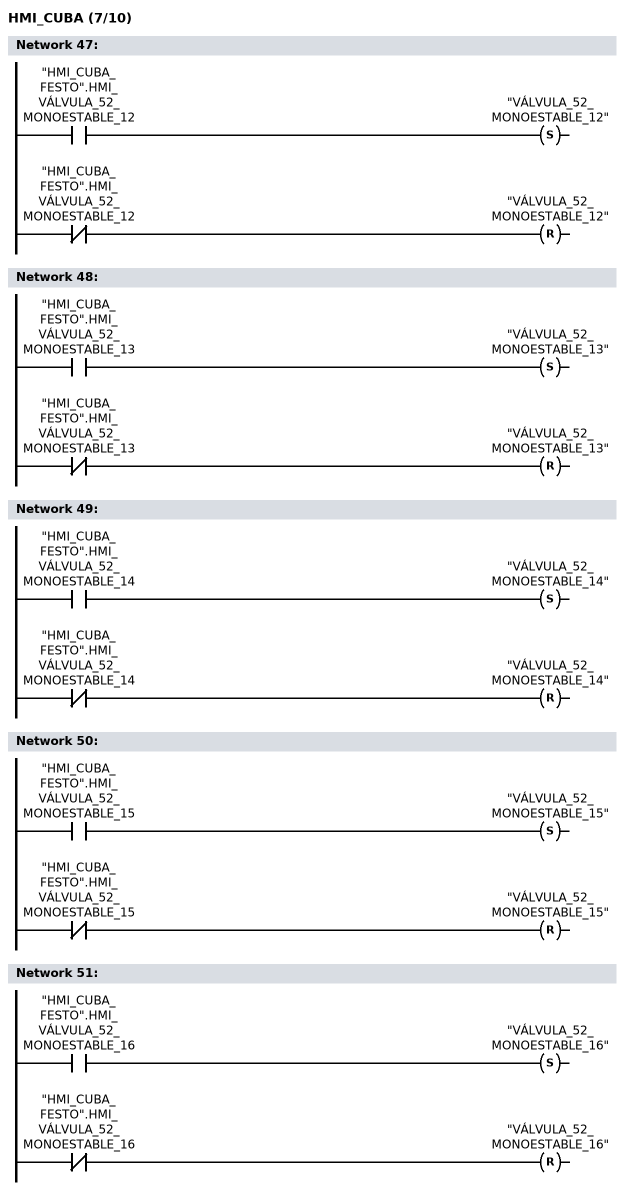
   RUNG wire#powerrail
      Contact( "HMI_CUBA_FESTO".HMI_VÁLVULA_52_MONOESTABLE_12 )
      S_Coil( "VÁLVULA_52_MONOESTABLE_12" )
   END_RUNG
   RUNG wire#powerrail
      I_Contact( "HMI_CUBA_FESTO".HMI_VÁLVULA_52_MONOESTABLE_12 )
      R_Coil( "VÁLVULA_52_MONOESTABLE_12" )
   END_RUNG
   // the same network as SCL:
   IF "HMI_CUBA_FESTO".HMI_VÁLVULA_52_MONOESTABLE_12 THEN "VÁLVULA_52_MONOESTABLE_12" := TRUE; END_IF;
   IF NOT "HMI_CUBA_FESTO".HMI_VÁLVULA_52_MONOESTABLE_12 THEN "VÁLVULA_52_MONOESTABLE_12" := FALSE; END_IF;
END_REGION

REGION Network 48
   RUNG wire#powerrail
      Contact( "HMI_CUBA_FESTO".HMI_VÁLVULA_52_MONOESTABLE_13 )
      S_Coil( "VÁLVULA_52_MONOESTABLE_13" )
   END_RUNG
   RUNG wire#powerrail
      I_Contact( "HMI_CUBA_FESTO".HMI_VÁLVULA_52_MONOESTABLE_13 )
      R_Coil( "VÁLVULA_52_MONOESTABLE_13" )
   END_RUNG
   // the same network as SCL:
   IF "HMI_CUBA_FESTO".HMI_VÁLVULA_52_MONOESTABLE_13 THEN "VÁLVULA_52_MONOESTABLE_13" := TRUE; END_IF;
   IF NOT "HMI_CUBA_FESTO".HMI_VÁLVULA_52_MONOESTABLE_13 THEN "VÁLVULA_52_MONOESTABLE_13" := FALSE; END_IF;
END_REGION

REGION Network 49
   RUNG wire#powerrail
      Contact( "HMI_CUBA_FESTO".HMI_VÁLVULA_52_MONOESTABLE_14 )
      S_Coil( "VÁLVULA_52_MONOESTABLE_14" )
   END_RUNG
   RUNG wire#powerrail
      I_Contact( "HMI_CUBA_FESTO".HMI_VÁLVULA_52_MONOESTABLE_14 )
      R_Coil( "VÁLVULA_52_MONOESTABLE_14" )
   END_RUNG
   // the same network as SCL:
   IF "HMI_CUBA_FESTO".HMI_VÁLVULA_52_MONOESTABLE_14 THEN "VÁLVULA_52_MONOESTABLE_14" := TRUE; END_IF;
   IF NOT "HMI_CUBA_FESTO".HMI_VÁLVULA_52_MONOESTABLE_14 THEN "VÁLVULA_52_MONOESTABLE_14" := FALSE; END_IF;
END_REGION

REGION Network 50
   RUNG wire#powerrail
      Contact( "HMI_CUBA_FESTO".HMI_VÁLVULA_52_MONOESTABLE_15 )
      S_Coil( "VÁLVULA_52_MONOESTABLE_15" )
   END_RUNG
   RUNG wire#powerrail
      I_Contact( "HMI_CUBA_FESTO".HMI_VÁLVULA_52_MONOESTABLE_15 )
      R_Coil( "VÁLVULA_52_MONOESTABLE_15" )
   END_RUNG
   // the same network as SCL:
   IF "HMI_CUBA_FESTO".HMI_VÁLVULA_52_MONOESTABLE_15 THEN "VÁLVULA_52_MONOESTABLE_15" := TRUE; END_IF;
   IF NOT "HMI_CUBA_FESTO".HMI_VÁLVULA_52_MONOESTABLE_15 THEN "VÁLVULA_52_MONOESTABLE_15" := FALSE; END_IF;
END_REGION

REGION Network 51
   RUNG wire#powerrail
      Contact( "HMI_CUBA_FESTO".HMI_VÁLVULA_52_MONOESTABLE_16 )
      S_Coil( "VÁLVULA_52_MONOESTABLE_16" )
   END_RUNG
   RUNG wire#powerrail
      I_Contact( "HMI_CUBA_FESTO".HMI_VÁLVULA_52_MONOESTABLE_16 )
      R_Coil( "VÁLVULA_52_MONOESTABLE_16" )
   END_RUNG
   // the same network as SCL:
   IF "HMI_CUBA_FESTO".HMI_VÁLVULA_52_MONOESTABLE_16 THEN "VÁLVULA_52_MONOESTABLE_16" := TRUE; END_IF;
   IF NOT "HMI_CUBA_FESTO".HMI_VÁLVULA_52_MONOESTABLE_16 THEN "VÁLVULA_52_MONOESTABLE_16" := FALSE; END_IF;
END_REGION

REGION Network 52
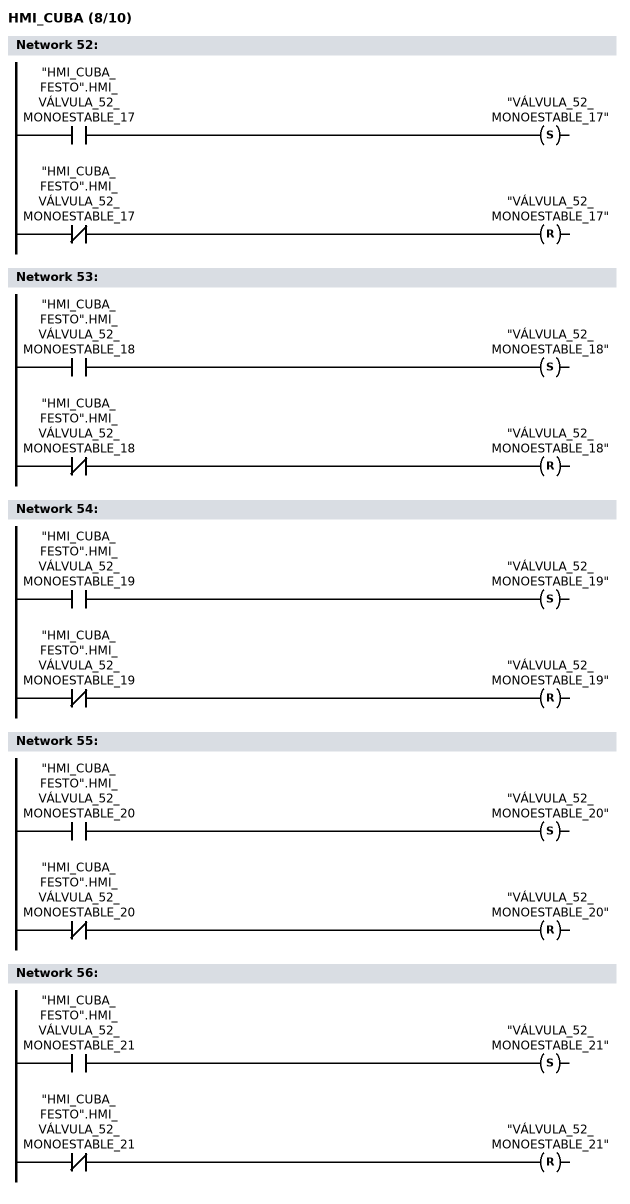
   RUNG wire#powerrail
      Contact( "HMI_CUBA_FESTO".HMI_VÁLVULA_52_MONOESTABLE_17 )
      S_Coil( "VÁLVULA_52_MONOESTABLE_17" )
   END_RUNG
   RUNG wire#powerrail
      I_Contact( "HMI_CUBA_FESTO".HMI_VÁLVULA_52_MONOESTABLE_17 )
      R_Coil( "VÁLVULA_52_MONOESTABLE_17" )
   END_RUNG
   // the same network as SCL:
   IF "HMI_CUBA_FESTO".HMI_VÁLVULA_52_MONOESTABLE_17 THEN "VÁLVULA_52_MONOESTABLE_17" := TRUE; END_IF;
   IF NOT "HMI_CUBA_FESTO".HMI_VÁLVULA_52_MONOESTABLE_17 THEN "VÁLVULA_52_MONOESTABLE_17" := FALSE; END_IF;
END_REGION

REGION Network 53
   RUNG wire#powerrail
      Contact( "HMI_CUBA_FESTO".HMI_VÁLVULA_52_MONOESTABLE_18 )
      S_Coil( "VÁLVULA_52_MONOESTABLE_18" )
   END_RUNG
   RUNG wire#powerrail
      I_Contact( "HMI_CUBA_FESTO".HMI_VÁLVULA_52_MONOESTABLE_18 )
      R_Coil( "VÁLVULA_52_MONOESTABLE_18" )
   END_RUNG
   // the same network as SCL:
   IF "HMI_CUBA_FESTO".HMI_VÁLVULA_52_MONOESTABLE_18 THEN "VÁLVULA_52_MONOESTABLE_18" := TRUE; END_IF;
   IF NOT "HMI_CUBA_FESTO".HMI_VÁLVULA_52_MONOESTABLE_18 THEN "VÁLVULA_52_MONOESTABLE_18" := FALSE; END_IF;
END_REGION

REGION Network 54
   RUNG wire#powerrail
      Contact( "HMI_CUBA_FESTO".HMI_VÁLVULA_52_MONOESTABLE_19 )
      S_Coil( "VÁLVULA_52_MONOESTABLE_19" )
   END_RUNG
   RUNG wire#powerrail
      I_Contact( "HMI_CUBA_FESTO".HMI_VÁLVULA_52_MONOESTABLE_19 )
      R_Coil( "VÁLVULA_52_MONOESTABLE_19" )
   END_RUNG
   // the same network as SCL:
   IF "HMI_CUBA_FESTO".HMI_VÁLVULA_52_MONOESTABLE_19 THEN "VÁLVULA_52_MONOESTABLE_19" := TRUE; END_IF;
   IF NOT "HMI_CUBA_FESTO".HMI_VÁLVULA_52_MONOESTABLE_19 THEN "VÁLVULA_52_MONOESTABLE_19" := FALSE; END_IF;
END_REGION

REGION Network 55
   RUNG wire#powerrail
      Contact( "HMI_CUBA_FESTO".HMI_VÁLVULA_52_MONOESTABLE_20 )
      S_Coil( "VÁLVULA_52_MONOESTABLE_20" )
   END_RUNG
   RUNG wire#powerrail
      I_Contact( "HMI_CUBA_FESTO".HMI_VÁLVULA_52_MONOESTABLE_20 )
      R_Coil( "VÁLVULA_52_MONOESTABLE_20" )
   END_RUNG
   // the same network as SCL:
   IF "HMI_CUBA_FESTO".HMI_VÁLVULA_52_MONOESTABLE_20 THEN "VÁLVULA_52_MONOESTABLE_20" := TRUE; END_IF;
   IF NOT "HMI_CUBA_FESTO".HMI_VÁLVULA_52_MONOESTABLE_20 THEN "VÁLVULA_52_MONOESTABLE_20" := FALSE; END_IF;
END_REGION

REGION Network 56
   RUNG wire#powerrail
      Contact( "HMI_CUBA_FESTO".HMI_VÁLVULA_52_MONOESTABLE_21 )
      S_Coil( "VÁLVULA_52_MONOESTABLE_21" )
   END_RUNG
   RUNG wire#powerrail
      I_Contact( "HMI_CUBA_FESTO".HMI_VÁLVULA_52_MONOESTABLE_21 )
      R_Coil( "VÁLVULA_52_MONOESTABLE_21" )
   END_RUNG
   // the same network as SCL:
   IF "HMI_CUBA_FESTO".HMI_VÁLVULA_52_MONOESTABLE_21 THEN "VÁLVULA_52_MONOESTABLE_21" := TRUE; END_IF;
   IF NOT "HMI_CUBA_FESTO".HMI_VÁLVULA_52_MONOESTABLE_21 THEN "VÁLVULA_52_MONOESTABLE_21" := FALSE; END_IF;
END_REGION

REGION Network 57
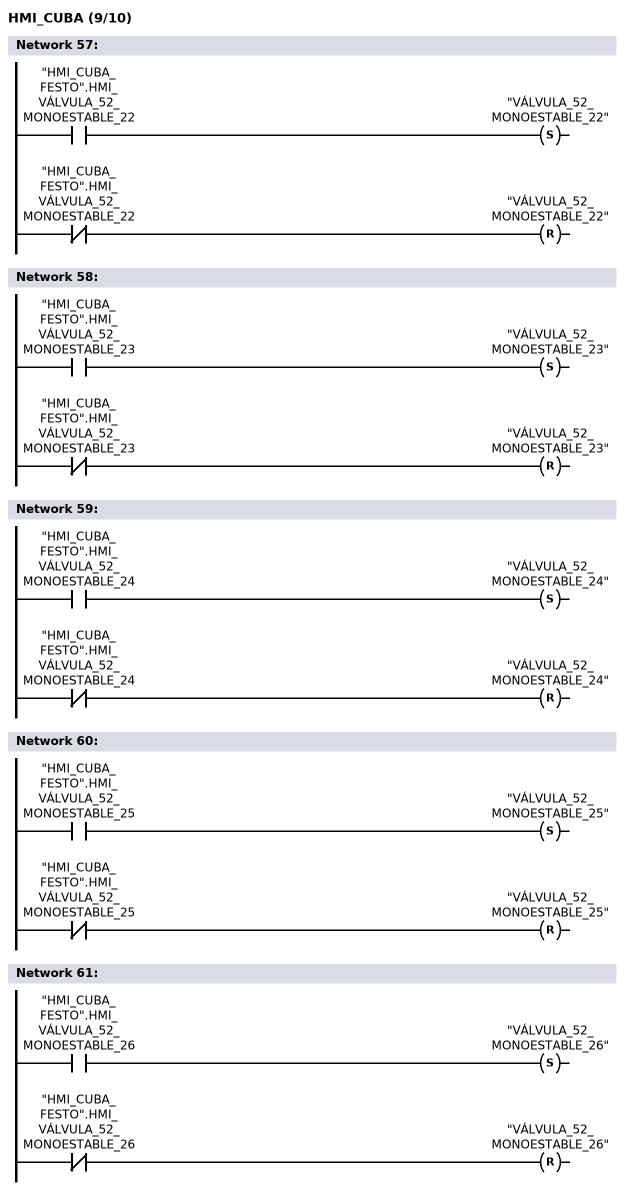
   RUNG wire#powerrail
      Contact( "HMI_CUBA_FESTO".HMI_VÁLVULA_52_MONOESTABLE_22 )
      S_Coil( "VÁLVULA_52_MONOESTABLE_22" )
   END_RUNG
   RUNG wire#powerrail
      I_Contact( "HMI_CUBA_FESTO".HMI_VÁLVULA_52_MONOESTABLE_22 )
      R_Coil( "VÁLVULA_52_MONOESTABLE_22" )
   END_RUNG
   // the same network as SCL:
   IF "HMI_CUBA_FESTO".HMI_VÁLVULA_52_MONOESTABLE_22 THEN "VÁLVULA_52_MONOESTABLE_22" := TRUE; END_IF;
   IF NOT "HMI_CUBA_FESTO".HMI_VÁLVULA_52_MONOESTABLE_22 THEN "VÁLVULA_52_MONOESTABLE_22" := FALSE; END_IF;
END_REGION

REGION Network 58
   RUNG wire#powerrail
      Contact( "HMI_CUBA_FESTO".HMI_VÁLVULA_52_MONOESTABLE_23 )
      S_Coil( "VÁLVULA_52_MONOESTABLE_23" )
   END_RUNG
   RUNG wire#powerrail
      I_Contact( "HMI_CUBA_FESTO".HMI_VÁLVULA_52_MONOESTABLE_23 )
      R_Coil( "VÁLVULA_52_MONOESTABLE_23" )
   END_RUNG
   // the same network as SCL:
   IF "HMI_CUBA_FESTO".HMI_VÁLVULA_52_MONOESTABLE_23 THEN "VÁLVULA_52_MONOESTABLE_23" := TRUE; END_IF;
   IF NOT "HMI_CUBA_FESTO".HMI_VÁLVULA_52_MONOESTABLE_23 THEN "VÁLVULA_52_MONOESTABLE_23" := FALSE; END_IF;
END_REGION

REGION Network 59
   RUNG wire#powerrail
      Contact( "HMI_CUBA_FESTO".HMI_VÁLVULA_52_MONOESTABLE_24 )
      S_Coil( "VÁLVULA_52_MONOESTABLE_24" )
   END_RUNG
   RUNG wire#powerrail
      I_Contact( "HMI_CUBA_FESTO".HMI_VÁLVULA_52_MONOESTABLE_24 )
      R_Coil( "VÁLVULA_52_MONOESTABLE_24" )
   END_RUNG
   // the same network as SCL:
   IF "HMI_CUBA_FESTO".HMI_VÁLVULA_52_MONOESTABLE_24 THEN "VÁLVULA_52_MONOESTABLE_24" := TRUE; END_IF;
   IF NOT "HMI_CUBA_FESTO".HMI_VÁLVULA_52_MONOESTABLE_24 THEN "VÁLVULA_52_MONOESTABLE_24" := FALSE; END_IF;
END_REGION

REGION Network 60
   RUNG wire#powerrail
      Contact( "HMI_CUBA_FESTO".HMI_VÁLVULA_52_MONOESTABLE_25 )
      S_Coil( "VÁLVULA_52_MONOESTABLE_25" )
   END_RUNG
   RUNG wire#powerrail
      I_Contact( "HMI_CUBA_FESTO".HMI_VÁLVULA_52_MONOESTABLE_25 )
      R_Coil( "VÁLVULA_52_MONOESTABLE_25" )
   END_RUNG
   // the same network as SCL:
   IF "HMI_CUBA_FESTO".HMI_VÁLVULA_52_MONOESTABLE_25 THEN "VÁLVULA_52_MONOESTABLE_25" := TRUE; END_IF;
   IF NOT "HMI_CUBA_FESTO".HMI_VÁLVULA_52_MONOESTABLE_25 THEN "VÁLVULA_52_MONOESTABLE_25" := FALSE; END_IF;
END_REGION

REGION Network 61
   RUNG wire#powerrail
      Contact( "HMI_CUBA_FESTO".HMI_VÁLVULA_52_MONOESTABLE_26 )
      S_Coil( "VÁLVULA_52_MONOESTABLE_26" )
   END_RUNG
   RUNG wire#powerrail
      I_Contact( "HMI_CUBA_FESTO".HMI_VÁLVULA_52_MONOESTABLE_26 )
      R_Coil( "VÁLVULA_52_MONOESTABLE_26" )
   END_RUNG
   // the same network as SCL:
   IF "HMI_CUBA_FESTO".HMI_VÁLVULA_52_MONOESTABLE_26 THEN "VÁLVULA_52_MONOESTABLE_26" := TRUE; END_IF;
   IF NOT "HMI_CUBA_FESTO".HMI_VÁLVULA_52_MONOESTABLE_26 THEN "VÁLVULA_52_MONOESTABLE_26" := FALSE; END_IF;
END_REGION

REGION Network 62
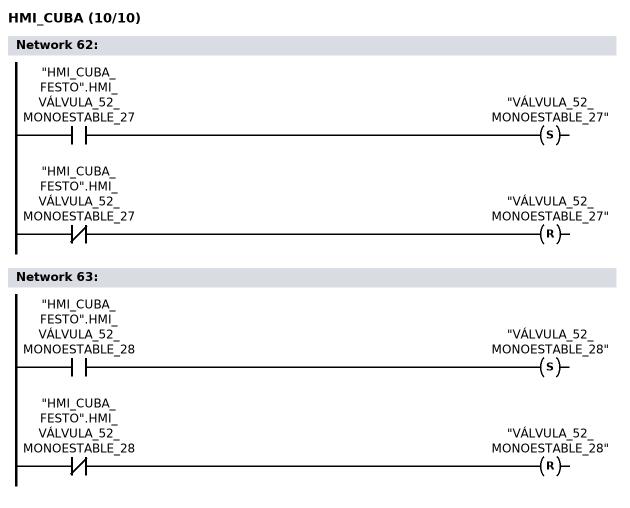
   RUNG wire#powerrail
      Contact( "HMI_CUBA_FESTO".HMI_VÁLVULA_52_MONOESTABLE_27 )
      S_Coil( "VÁLVULA_52_MONOESTABLE_27" )
   END_RUNG
   RUNG wire#powerrail
      I_Contact( "HMI_CUBA_FESTO".HMI_VÁLVULA_52_MONOESTABLE_27 )
      R_Coil( "VÁLVULA_52_MONOESTABLE_27" )
   END_RUNG
   // the same network as SCL:
   IF "HMI_CUBA_FESTO".HMI_VÁLVULA_52_MONOESTABLE_27 THEN "VÁLVULA_52_MONOESTABLE_27" := TRUE; END_IF;
   IF NOT "HMI_CUBA_FESTO".HMI_VÁLVULA_52_MONOESTABLE_27 THEN "VÁLVULA_52_MONOESTABLE_27" := FALSE; END_IF;
END_REGION

REGION Network 63
   RUNG wire#powerrail
      Contact( "HMI_CUBA_FESTO".HMI_VÁLVULA_52_MONOESTABLE_28 )
      S_Coil( "VÁLVULA_52_MONOESTABLE_28" )
   END_RUNG
   RUNG wire#powerrail
      I_Contact( "HMI_CUBA_FESTO".HMI_VÁLVULA_52_MONOESTABLE_28 )
      R_Coil( "VÁLVULA_52_MONOESTABLE_28" )
   END_RUNG
   // the same network as SCL:
   IF "HMI_CUBA_FESTO".HMI_VÁLVULA_52_MONOESTABLE_28 THEN "VÁLVULA_52_MONOESTABLE_28" := TRUE; END_IF;
   IF NOT "HMI_CUBA_FESTO".HMI_VÁLVULA_52_MONOESTABLE_28 THEN "VÁLVULA_52_MONOESTABLE_28" := FALSE; END_IF;
END_REGION
END_FUNCTION_BLOCK

FUNCTION_BLOCK "GIRO_POSITIVO"   // FB10, LAD
{ S7_Optimized_Access := 'TRUE' }
VERSION : 0.1
   VAR_TEMP   // added for the SCL form of the ladder/FBD networks
      _w1 : Bool;
   END_VAR
BEGIN

REGION Network 1: Estado 1
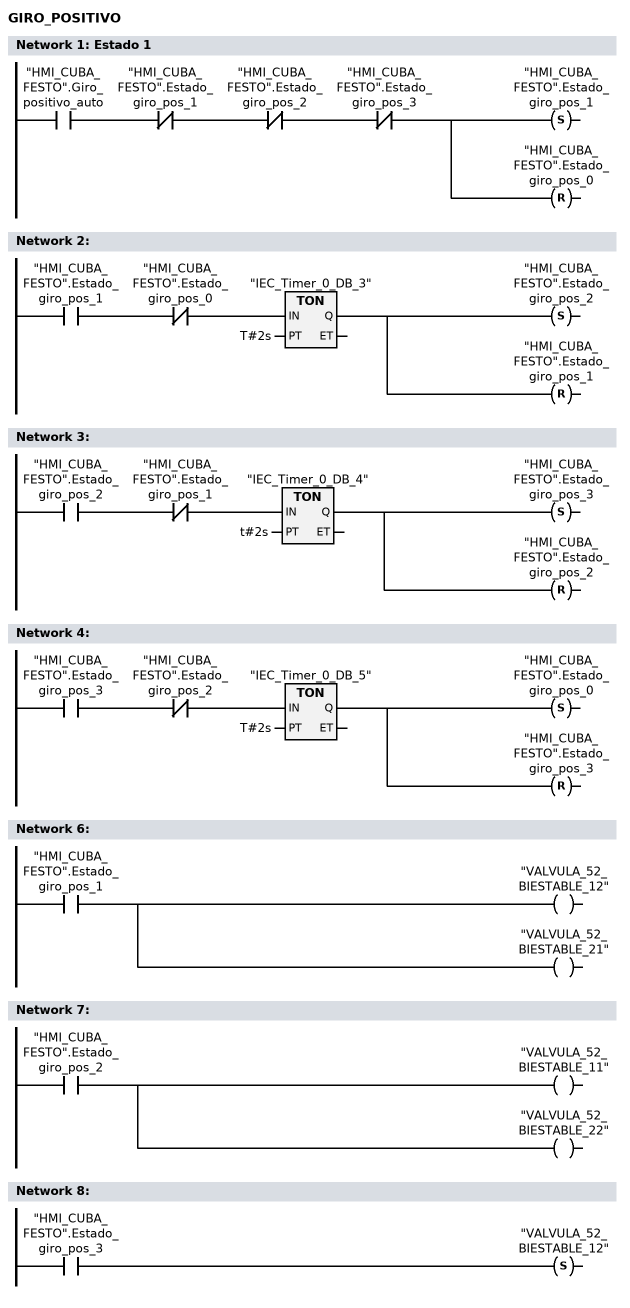
   RUNG wire#powerrail
      Contact( "HMI_CUBA_FESTO".Giro_positivo_auto )
      I_Contact( "HMI_CUBA_FESTO".Estado_giro_pos_1 )
      I_Contact( "HMI_CUBA_FESTO".Estado_giro_pos_2 )
      I_Contact( "HMI_CUBA_FESTO".Estado_giro_pos_3 )
      wire#w1
      S_Coil( "HMI_CUBA_FESTO".Estado_giro_pos_1 )
   END_RUNG
   RUNG wire#w1
      R_Coil( "HMI_CUBA_FESTO".Estado_giro_pos_0 )
   END_RUNG
   // the same network as SCL:
   #_w1 := "HMI_CUBA_FESTO".Giro_positivo_auto AND NOT "HMI_CUBA_FESTO".Estado_giro_pos_1 AND NOT "HMI_CUBA_FESTO".Estado_giro_pos_2 AND NOT "HMI_CUBA_FESTO".Estado_giro_pos_3;
   IF #_w1 THEN
       "HMI_CUBA_FESTO".Estado_giro_pos_1 := TRUE;
       "HMI_CUBA_FESTO".Estado_giro_pos_0 := FALSE;
   END_IF;
END_REGION

REGION Network 2
   "IEC_Timer_0_DB_3".TON(IN := "HMI_CUBA_FESTO".Estado_giro_pos_1 AND NOT "HMI_CUBA_FESTO".Estado_giro_pos_0,
                          PT := T#2s);
   IF "IEC_Timer_0_DB_3".Q THEN
       "HMI_CUBA_FESTO".Estado_giro_pos_2 := TRUE;
       "HMI_CUBA_FESTO".Estado_giro_pos_1 := FALSE;
   END_IF;
END_REGION

REGION Network 3
   "IEC_Timer_0_DB_4".TON(IN := "HMI_CUBA_FESTO".Estado_giro_pos_2 AND NOT "HMI_CUBA_FESTO".Estado_giro_pos_1,
                          PT := t#2s);
   IF "IEC_Timer_0_DB_4".Q THEN
       "HMI_CUBA_FESTO".Estado_giro_pos_3 := TRUE;
       "HMI_CUBA_FESTO".Estado_giro_pos_2 := FALSE;
   END_IF;
END_REGION

REGION Network 4
   "IEC_Timer_0_DB_5".TON(IN := "HMI_CUBA_FESTO".Estado_giro_pos_3 AND NOT "HMI_CUBA_FESTO".Estado_giro_pos_2,
                          PT := T#2s);
   IF "IEC_Timer_0_DB_5".Q THEN
       "HMI_CUBA_FESTO".Estado_giro_pos_0 := TRUE;
       "HMI_CUBA_FESTO".Estado_giro_pos_3 := FALSE;
   END_IF;
END_REGION

REGION Network 6
   RUNG wire#powerrail
      Contact( "HMI_CUBA_FESTO".Estado_giro_pos_1 )
      wire#w1
      Coil( "VALVULA_52_BIESTABLE_12" )
   END_RUNG
   RUNG wire#w1
      Coil( "VALVULA_52_BIESTABLE_21" )
   END_RUNG
   // the same network as SCL:
   "VALVULA_52_BIESTABLE_12" := "HMI_CUBA_FESTO".Estado_giro_pos_1;
   "VALVULA_52_BIESTABLE_21" := "HMI_CUBA_FESTO".Estado_giro_pos_1;
END_REGION

REGION Network 7
   RUNG wire#powerrail
      Contact( "HMI_CUBA_FESTO".Estado_giro_pos_2 )
      wire#w1
      Coil( "VALVULA_52_BIESTABLE_11" )
   END_RUNG
   RUNG wire#w1
      Coil( "VALVULA_52_BIESTABLE_22" )
   END_RUNG
   // the same network as SCL:
   "VALVULA_52_BIESTABLE_11" := "HMI_CUBA_FESTO".Estado_giro_pos_2;
   "VALVULA_52_BIESTABLE_22" := "HMI_CUBA_FESTO".Estado_giro_pos_2;
END_REGION

REGION Network 8
   RUNG wire#powerrail
      Contact( "HMI_CUBA_FESTO".Estado_giro_pos_3 )
      S_Coil( "VALVULA_52_BIESTABLE_12" )
   END_RUNG
   // the same network as SCL:
   IF "HMI_CUBA_FESTO".Estado_giro_pos_3 THEN "VALVULA_52_BIESTABLE_12" := TRUE; END_IF;
END_REGION
END_FUNCTION_BLOCK

FUNCTION_BLOCK "GIRO_NEGATIVO_1"   // FB14, LAD
{ S7_Optimized_Access := 'TRUE' }
VERSION : 0.1
   VAR_TEMP   // added for the SCL form of the ladder/FBD networks
      _w1 : Bool;
   END_VAR
BEGIN

REGION Network 1: Estado 1
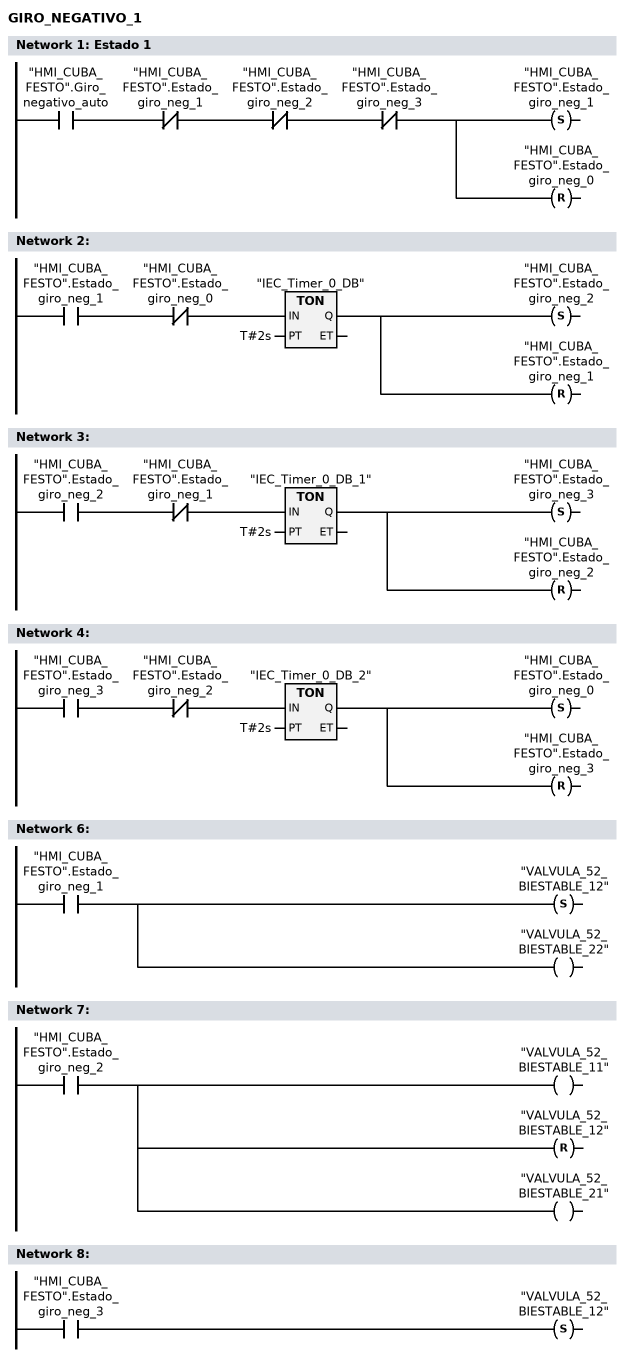
   RUNG wire#powerrail
      Contact( "HMI_CUBA_FESTO".Giro_negativo_auto )
      I_Contact( "HMI_CUBA_FESTO".Estado_giro_neg_1 )
      I_Contact( "HMI_CUBA_FESTO".Estado_giro_neg_2 )
      I_Contact( "HMI_CUBA_FESTO".Estado_giro_neg_3 )
      wire#w1
      S_Coil( "HMI_CUBA_FESTO".Estado_giro_neg_1 )
   END_RUNG
   RUNG wire#w1
      R_Coil( "HMI_CUBA_FESTO".Estado_giro_neg_0 )
   END_RUNG
   // the same network as SCL:
   #_w1 := "HMI_CUBA_FESTO".Giro_negativo_auto AND NOT "HMI_CUBA_FESTO".Estado_giro_neg_1 AND NOT "HMI_CUBA_FESTO".Estado_giro_neg_2 AND NOT "HMI_CUBA_FESTO".Estado_giro_neg_3;
   IF #_w1 THEN
       "HMI_CUBA_FESTO".Estado_giro_neg_1 := TRUE;
       "HMI_CUBA_FESTO".Estado_giro_neg_0 := FALSE;
   END_IF;
END_REGION

REGION Network 2
   "IEC_Timer_0_DB".TON(IN := "HMI_CUBA_FESTO".Estado_giro_neg_1 AND NOT "HMI_CUBA_FESTO".Estado_giro_neg_0,
                        PT := T#2s);
   IF "IEC_Timer_0_DB".Q THEN
       "HMI_CUBA_FESTO".Estado_giro_neg_2 := TRUE;
       "HMI_CUBA_FESTO".Estado_giro_neg_1 := FALSE;
   END_IF;
END_REGION

REGION Network 3
   "IEC_Timer_0_DB_1".TON(IN := "HMI_CUBA_FESTO".Estado_giro_neg_2 AND NOT "HMI_CUBA_FESTO".Estado_giro_neg_1,
                          PT := T#2s);
   IF "IEC_Timer_0_DB_1".Q THEN
       "HMI_CUBA_FESTO".Estado_giro_neg_3 := TRUE;
       "HMI_CUBA_FESTO".Estado_giro_neg_2 := FALSE;
   END_IF;
END_REGION

REGION Network 4
   "IEC_Timer_0_DB_2".TON(IN := "HMI_CUBA_FESTO".Estado_giro_neg_3 AND NOT "HMI_CUBA_FESTO".Estado_giro_neg_2,
                          PT := T#2s);
   IF "IEC_Timer_0_DB_2".Q THEN
       "HMI_CUBA_FESTO".Estado_giro_neg_0 := TRUE;
       "HMI_CUBA_FESTO".Estado_giro_neg_3 := FALSE;
   END_IF;
END_REGION

REGION Network 6
   RUNG wire#powerrail
      Contact( "HMI_CUBA_FESTO".Estado_giro_neg_1 )
      wire#w1
      S_Coil( "VALVULA_52_BIESTABLE_12" )
   END_RUNG
   RUNG wire#w1
      Coil( "VALVULA_52_BIESTABLE_22" )
   END_RUNG
   // the same network as SCL:
   IF "HMI_CUBA_FESTO".Estado_giro_neg_1 THEN "VALVULA_52_BIESTABLE_12" := TRUE; END_IF;
   "VALVULA_52_BIESTABLE_22" := "HMI_CUBA_FESTO".Estado_giro_neg_1;
END_REGION

REGION Network 7
   RUNG wire#powerrail
      Contact( "HMI_CUBA_FESTO".Estado_giro_neg_2 )
      wire#w1
      Coil( "VALVULA_52_BIESTABLE_11" )
   END_RUNG
   RUNG wire#w1
      R_Coil( "VALVULA_52_BIESTABLE_12" )
   END_RUNG
   RUNG wire#w1
      Coil( "VALVULA_52_BIESTABLE_21" )
   END_RUNG
   // the same network as SCL:
   "VALVULA_52_BIESTABLE_11" := "HMI_CUBA_FESTO".Estado_giro_neg_2;
   IF "HMI_CUBA_FESTO".Estado_giro_neg_2 THEN "VALVULA_52_BIESTABLE_12" := FALSE; END_IF;
   "VALVULA_52_BIESTABLE_21" := "HMI_CUBA_FESTO".Estado_giro_neg_2;
END_REGION

REGION Network 8
   RUNG wire#powerrail
      Contact( "HMI_CUBA_FESTO".Estado_giro_neg_3 )
      S_Coil( "VALVULA_52_BIESTABLE_12" )
   END_RUNG
   // the same network as SCL:
   IF "HMI_CUBA_FESTO".Estado_giro_neg_3 THEN "VALVULA_52_BIESTABLE_12" := TRUE; END_IF;
END_REGION
END_FUNCTION_BLOCK

// folder: Achim

FUNCTION_BLOCK "Achim_testPepaFrk"   // FB8, LAD
TITLE = test tools
{ S7_Optimized_Access := 'TRUE' }
VERSION : 0.1
   VAR_INPUT
      inToolIdProxy1 : Bool;
      inToolIdProxy2 : Bool;
      inToolIdProxy3 : Bool;
      inToolIdProxy4 : Bool;
      inAirActivate : Bool;
      inAirPepaCylInActivate : Bool;
      inAirPepaCylOutActivate : Bool;
      inWaterInspPumpActivate : Bool;
      inWaterActivate : Bool;
      inStopRobot : Bool;
      inContRobot : Bool;
      inResetAlarms : Bool;
      inInspRunning : Bool;
      inSTOPMESS : Bool;
      inPRO_ACT : Bool;
      inWaterInspPumpRunning : Bool;
      inWaterInspAlarmFilter : Bool;
      inWaterInspAlarmFc : Bool;
      inWaterInspAlarmElecProt : Bool;
      inWaterInspAlarmUv : Bool;
      inWaterInspAlarmLowLevel : Bool;
      inPepaCylInProxy : Bool;
      inPepaCylOutProxy : Bool;
      inAirOprProxy : Bool;
      inAirMpsCoupledE1 : Bool;
      inAirMpsLockedE2 : Bool;
      inAirMpsUnlockedE3 : Bool;
      inAirMpsPressD1 : Bool;
      inFrkLs1Nc1 : Bool;
      inFrkLs1Nc2 : Bool;
      inFrkLs2Nc1 : Bool;
      inFrkLs2Nc2 : Bool;
      airMpsTimeout : Time := T#500ms;
      airPepaCylTimeout : Time := T#100ms;
      frkLsTimeout : Time := T#100ms;
   END_VAR
   VAR_OUTPUT
      outWaterInspEvL1 : Bool;
      outWaterInspEvL2 : Bool;
      outWaterInspPanelS1 : Bool;
      outWaterInspPanelS2 : Bool;
      outWaterInspPanelS3 : Bool;
      outWaterInspPump : Bool;
      outAirEvOpr : Bool;
      outAirEvMps : Bool;
      outAirPepaCylIn : Bool;
      outAirPepaCylOut : Bool;
      outAntiSpash1 : Bool;
      outAntiSpash2 : Bool;
      outAirMpsAlarm : Bool;
      outAirOprAlarm : Bool;
      outPepaCylAlarm : Bool;
      outFrkLsAlarm : Bool;
      outWaterInspAlarm : Bool;
      outWaterInspAdv : Bool;
      outStopRobot : Bool;
      outMOVE_ENABLE : Bool;
      outCONF_MESS : Bool;
      outEXT_START : Bool;
   END_VAR
   VAR
      tonMpsOn : TON_TIME;
      tonPepaCylOut : TON_TIME;
      tonFrkLs : TON_TIME;
      staticStoppingAlarm : Bool;
      staticAirMpsAlarm : Bool;
      staticAirOprAlarm : Bool;
      staticPepaCylAlarm : Bool;
      staticFrkLsAlarm : Bool;
      staticWaterInspAlarm : Bool;
      staticWaterInspAdv : Bool;
      staticStopRobot : Bool;
      staticContRobot : Bool;
      staticRobotWasStopped : Bool;
      staticairMpsOk : Bool;
      staticTool : Int;
      rtStopRobot : R_TRIG;
      rtContRobot : R_TRIG;
   END_VAR
BEGIN

REGION Network 1 (SCL)
   // tool identification
   IF #inToolIdProxy1 AND NOT #inToolIdProxy2 AND NOT #inToolIdProxy3 AND NOT #inToolIdProxy4 THEN
       #staticTool := 1; // PEPA
   ELSIF NOT #inToolIdProxy1 AND #inToolIdProxy2 AND NOT #inToolIdProxy3 AND NOT #inToolIdProxy4 THEN
       #staticTool := 2; // pole
   ELSIF #inToolIdProxy1 AND #inToolIdProxy2 AND NOT #inToolIdProxy3 AND NOT #inToolIdProxy4 THEN
       #staticTool := 3; // fork
   ELSIF NOT #inToolIdProxy1 AND NOT #inToolIdProxy2 AND #inToolIdProxy3 AND NOT #inToolIdProxy4 THEN
       #staticTool := 4; // teaching
   ELSIF #inToolIdProxy1 AND NOT #inToolIdProxy2 AND #inToolIdProxy3 AND NOT #inToolIdProxy4 THEN
       #staticTool := 5; // marker    
   ELSIF NOT #inToolIdProxy1 AND NOT #inToolIdProxy2 AND NOT #inToolIdProxy3 AND NOT #inToolIdProxy4 THEN
       #staticTool := 0; // no tool  
   ELSE
       #staticTool := -1; // unknown
   END_IF;

   // air MPS & OPR activation
   #outAirEvOpr := #inAirActivate AND (#staticTool=1 OR #staticTool=2 OR #staticTool=5);
   #outAirEvMps := #inAirActivate;

   // check MPS & OPR signals
   #staticairMpsOk := #inAirMpsCoupledE1 AND #inAirMpsLockedE2 AND NOT #inAirMpsUnlockedE3 AND #inAirMpsPressD1;
   #tonMpsOn(IN := #inAirActivate AND #staticTool>0,
                 PT := #airMpsTimeout);
   IF #tonMpsOn.Q THEN
           IF NOT #staticairMpsOk THEN
               #staticAirMpsAlarm := true;
           END_IF;
           IF NOT #inAirOprProxy AND (#staticTool=1 OR #staticTool=2 OR #staticTool=5) THEN
               #staticAirOprAlarm := true;
           END_IF;
   END_IF;

   // alarms
   IF #inResetAlarms THEN
       #staticAirMpsAlarm := false;
       #staticAirOprAlarm := false;
       #staticPepaCylAlarm := false;
       #staticFrkLsAlarm := false;
       #staticWaterInspAlarm := false;
       #staticWaterInspAdv := false;
   END_IF;
   IF #inResetAlarms AND #inSTOPMESS THEN
       #outCONF_MESS := true;
   ELSE
       #outCONF_MESS := false;
   END_IF;

   #rtContRobot(CLK := #inContRobot);
   IF #staticRobotWasStopped AND #rtContRobot.Q AND NOT #staticStoppingAlarm THEN
       #staticContRobot := true;
       #staticRobotWasStopped := false;
   END_IF;

   // water pump
   IF #inWaterInspAlarmFilter OR #inWaterInspAlarmUv THEN
       #staticWaterInspAdv := true;
   END_IF;
   IF (#inWaterInspAlarmFc OR #inWaterInspAlarmElecProt OR #inWaterInspAlarmLowLevel) AND #inWaterActivate THEN
       #staticWaterInspAlarm := true;
   END_IF;
   #outWaterInspPump := #inWaterInspPumpActivate AND NOT #staticWaterInspAlarm;

   // water valves
   #outWaterInspPanelS1 := #inWaterActivate AND #inWaterInspPumpRunning AND #staticTool=3;
   #outWaterInspPanelS2 := #inWaterActivate AND #inWaterInspPumpRunning AND #staticTool=3;
   #outWaterInspPanelS3 := #inWaterActivate AND #inWaterInspPumpRunning AND #staticTool=1;
   #outWaterInspEvL1 := #inWaterActivate AND #inWaterInspPumpRunning AND #staticTool = 3;
   #outWaterInspEvL2 := #inWaterActivate AND #inWaterInspPumpRunning AND (#staticTool=1 OR #staticTool=3);

   // retract & extend PEPA / marker cylinder
   #outAirPepaCylIn := #inAirPepaCylInActivate AND (#staticTool=1 OR #staticTool=5);
   #outAirPepaCylOut := #inAirPepaCylOutActivate AND (#staticTool=1 OR #staticTool=5);

   // anti splash air FRK
   #outAntiSpash1 := #inInspRunning AND #staticTool=3;
   #outAntiSpash2 := #inInspRunning AND #staticTool=3;

   // check micro cyl in / cyl out triggers while PEPA cyl out during inspection
   #tonPepaCylOut(IN := #inInspRunning AND (#inPepaCylInProxy OR #inPepaCylOutProxy) AND (#staticTool=1 OR #staticTool=5),
                       PT := #airPepaCylTimeout);
   IF #tonPepaCylOut.Q THEN
       #staticPepaCylAlarm := true;
   END_IF;

   // check limit switches FRK
   #tonFrkLs(IN := (NOT #inFrkLs1Nc1 OR NOT #inFrkLs1Nc2 OR NOT #inFrkLs2Nc1 OR NOT #inFrkLs2Nc1 OR NOT #inFrkLs2Nc2) AND #staticTool=3,
             PT := #frkLsTimeout);
   IF #tonFrkLs.Q THEN
       #staticFrkLsAlarm := true;
   END_IF;

   // stop robot
   #staticStoppingAlarm := #staticAirMpsAlarm OR #staticAirOprAlarm OR #staticWaterInspAlarm OR #staticPepaCylAlarm OR #staticFrkLsAlarm;
   #rtStopRobot(CLK := #inStopRobot OR #staticStoppingAlarm);
   IF #rtStopRobot.Q THEN
       #staticStopRobot := true;
   END_IF;

   // feedback stop robot cmd from robot
   IF #staticStopRobot AND #inSTOPMESS AND NOT #inPRO_ACT THEN
       #staticStopRobot := false;
       #staticRobotWasStopped := true;
   END_IF;

   // feedback cont robot cmd from robot
   IF #staticContRobot AND #inPRO_ACT THEN
       #staticContRobot := false;
   END_IF;

   // outputs
   #outStopRobot := #staticStopRobot;
   #outMOVE_ENABLE := NOT #staticStopRobot;
   #outEXT_START := #staticContRobot;
   #outAirMpsAlarm := #staticAirMpsAlarm;
   #outAirOprAlarm := #staticAirOprAlarm;
   #outPepaCylAlarm := #staticPepaCylAlarm;
   #outFrkLsAlarm := #staticFrkLsAlarm;
   #outWaterInspAlarm := #staticWaterInspAlarm;
   #outWaterInspAdv := #staticWaterInspAdv;
END_REGION
END_FUNCTION_BLOCK

FUNCTION "Achim" : Void   // FC1, LAD
{ S7_Optimized_Access := 'TRUE' }
VERSION : 0.1
BEGIN

REGION Network 1: test end effector
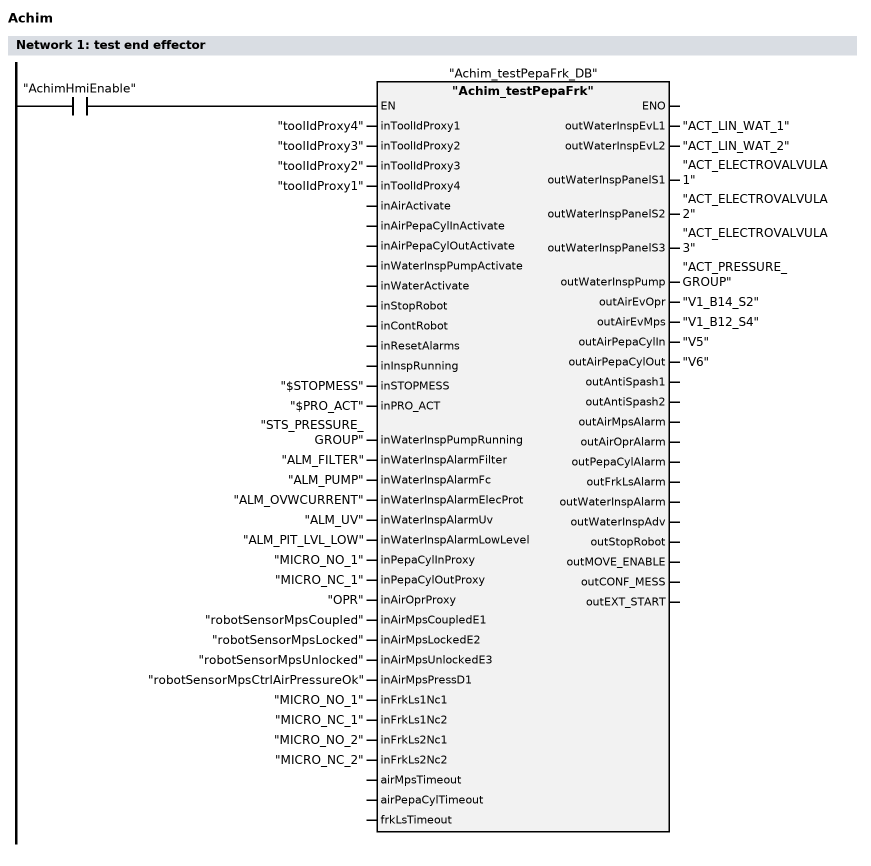
   RUNG wire#powerrail
      Contact( "AchimHmiEnable" )
      "Achim_testPepaFrk_DB"(inToolIdProxy1 := "toolIdProxy4", inToolIdProxy2 := "toolIdProxy3", inToolIdProxy3 := "toolIdProxy2", inToolIdProxy4 := "toolIdProxy1", inAirActivate :=, inAirPepaCylInActivate :=, inAirPepaCylOutActivate :=, inWaterInspPumpActivate :=, inWaterActivate :=, inStopRobot :=, inContRobot :=, inResetAlarms :=, inInspRunning :=, inSTOPMESS := "$STOPMESS", inPRO_ACT := "$PRO_ACT", inWaterInspPumpRunning := "STS_PRESSURE_GROUP", inWaterInspAlarmFilter := "ALM_FILTER", inWaterInspAlarmFc := "ALM_PUMP", inWaterInspAlarmElecProt := "ALM_OVWCURRENT", inWaterInspAlarmUv := "ALM_UV", inWaterInspAlarmLowLevel := "ALM_PIT_LVL_LOW", inPepaCylInProxy := "MICRO_NO_1", inPepaCylOutProxy := "MICRO_NC_1", inAirOprProxy := "OPR", inAirMpsCoupledE1 := "robotSensorMpsCoupled", inAirMpsLockedE2 := "robotSensorMpsLocked", inAirMpsUnlockedE3 := "robotSensorMpsUnlocked", inAirMpsPressD1 := "robotSensorMpsCtrlAirPressureOk", inFrkLs1Nc1 := "MICRO_NO_1", inFrkLs1Nc2 := "MICRO_NC_1", inFrkLs2Nc1 := "MICRO_NO_2", inFrkLs2Nc2 := "MICRO_NC_2", airMpsTimeout :=, airPepaCylTimeout :=, frkLsTimeout :=, outWaterInspEvL1 => "ACT_LIN_WAT_1", outWaterInspEvL2 => "ACT_LIN_WAT_2", outWaterInspPanelS1 => "ACT_ELECTROVALVULA1", outWaterInspPanelS2 => "ACT_ELECTROVALVULA2", outWaterInspPanelS3 => "ACT_ELECTROVALVULA3", outWaterInspPump => "ACT_PRESSURE_GROUP", outAirEvOpr => "V1_B14_S2", outAirEvMps => "V1_B12_S4", outAirPepaCylIn => "V5", outAirPepaCylOut => "V6", outAntiSpash1 =>, outAntiSpash2 =>, outAirMpsAlarm =>, outAirOprAlarm =>, outPepaCylAlarm =>, outFrkLsAlarm =>, outWaterInspAlarm =>, outWaterInspAdv =>, outStopRobot =>, outMOVE_ENABLE =>, outCONF_MESS =>, outEXT_START =>)
   END_RUNG
   // the same network as SCL:
   IF "AchimHmiEnable" THEN
       "Achim_testPepaFrk_DB"(inToolIdProxy1 := "toolIdProxy4",   // "Achim_testPepaFrk"
                              inToolIdProxy2 := "toolIdProxy3",
                              inToolIdProxy3 := "toolIdProxy2",
                              inToolIdProxy4 := "toolIdProxy1",
                              inSTOPMESS := "$STOPMESS",
                              inPRO_ACT := "$PRO_ACT",
                              inWaterInspPumpRunning := "STS_PRESSURE_GROUP",
                              inWaterInspAlarmFilter := "ALM_FILTER",
                              inWaterInspAlarmFc := "ALM_PUMP",
                              inWaterInspAlarmElecProt := "ALM_OVWCURRENT",
                              inWaterInspAlarmUv := "ALM_UV",
                              inWaterInspAlarmLowLevel := "ALM_PIT_LVL_LOW",
                              inPepaCylInProxy := "MICRO_NO_1",
                              inPepaCylOutProxy := "MICRO_NC_1",
                              inAirOprProxy := "OPR",
                              inAirMpsCoupledE1 := "robotSensorMpsCoupled",
                              inAirMpsLockedE2 := "robotSensorMpsLocked",
                              inAirMpsUnlockedE3 := "robotSensorMpsUnlocked",
                              inAirMpsPressD1 := "robotSensorMpsCtrlAirPressureOk",
                              inFrkLs1Nc1 := "MICRO_NO_1",
                              inFrkLs1Nc2 := "MICRO_NC_1",
                              inFrkLs2Nc1 := "MICRO_NO_2",
                              inFrkLs2Nc2 := "MICRO_NC_2",
                              outWaterInspEvL1 => "ACT_LIN_WAT_1",
                              outWaterInspEvL2 => "ACT_LIN_WAT_2",
                              outWaterInspPanelS1 => "ACT_ELECTROVALVULA1",
                              outWaterInspPanelS2 => "ACT_ELECTROVALVULA2",
                              outWaterInspPanelS3 => "ACT_ELECTROVALVULA3",
                              outWaterInspPump => "ACT_PRESSURE_GROUP",
                              outAirEvOpr => "V1_B14_S2",
                              outAirEvMps => "V1_B12_S4",
                              outAirPepaCylIn => "V5",
                              outAirPepaCylOut => "V6");
   END_IF;
END_REGION
END_FUNCTION

(* ===== HMI "HMI_RT_1" =====
system functions are stored by id; their names below are inferred from use
connection "HMI_Connection_1": ETHERNET, SMART_S7_1200_OMS

HMI tags "Default tag table"
   "Tag_ScreenNumber" : UInt, internal

HMI tags "CUBA_FESTO"
   "HMI_CUBA_FESTO_HMI_Sensor_plato_giro_1" : Bool = PLC HMI_CUBA_FESTO.HMI_Sensor_plato_giro_1, 100 ms
   "HMI_CUBA_FESTO_HMI_Sensor_Plato_giro_2" : Bool = PLC HMI_CUBA_FESTO.HMI_Sensor_Plato_giro_2, 100 ms
   "HMI_CUBA_FESTO_HMI_Sensor_plato_giro_3" : Bool = PLC HMI_CUBA_FESTO.HMI_Sensor_plato_giro_3, 100 ms
   "HMI_CUBA_FESTO_HMI_Sensor_ADN_bastidor_bloqueado_1" : Bool = PLC HMI_CUBA_FESTO.HMI_Sensor_ADN_bastidor_bloqueado_1, 100 ms
   "HMI_CUBA_FESTO_HMI_Sensor_ADN_bastidor_desbloqueado_1" : Bool = PLC HMI_CUBA_FESTO.HMI_Sensor_ADN_bastidor_desbloqueado_1, 100 ms
   "HMI_CUBA_FESTO_HMI_Sensor_ADN_bastidor_bloqueado_2" : Bool = PLC HMI_CUBA_FESTO.HMI_Sensor_ADN_bastidor_bloqueado_2, 100 ms
   "HMI_CUBA_FESTO_HMI_Sensor_ADN_bastidor_desbloqueado_2" : Bool = PLC HMI_CUBA_FESTO.HMI_Sensor_ADN_bastidor_desbloqueado_2, 100 ms
   "HMI_CUBA_FESTO_HMI_SENSOR_CRDSNU_BASTIDOR_BLOQUEADO_1" : Bool = PLC HMI_CUBA_FESTO.HMI_SENSOR_CRDSNU_BASTIDOR_BLOQUEADO_1, 100 ms
   "HMI_CUBA_FESTO_HMI_SENSOR_CRDSNU_BASTIDOR_DESBLOQUEADO_1" : Bool = PLC HMI_CUBA_FESTO.HMI_SENSOR_CRDSNU_BASTIDOR_DESBLOQUEADO_1, 100 ms
   "HMI_CUBA_FESTO_HMI_SENSOR_CRDSNU_BASTIDOR_BLOQUEADO_2" : Bool = PLC HMI_CUBA_FESTO.HMI_SENSOR_CRDSNU_BASTIDOR_BLOQUEADO_2, 100 ms
   "HMI_CUBA_FESTO_HMI_SENSOR_CRDSNU_BASTIDOR_DESBLOQUEADO_2" : Bool = PLC HMI_CUBA_FESTO.HMI_SENSOR_CRDSNU_BASTIDOR_DESBLOQUEADO_2, 100 ms
   "HMI_CUBA_FESTO_HMI_SENSOR_DSBG_BASTIDOR_ARRIBA_1" : Bool = PLC HMI_CUBA_FESTO.HMI_SENSOR_DSBG_BASTIDOR_ARRIBA_1, 100 ms
   "HMI_CUBA_FESTO_HMI_SENSOR_DSBG_BASTIDOR_ABAJO_1" : Bool = PLC HMI_CUBA_FESTO.HMI_SENSOR_DSBG_BASTIDOR_ABAJO_1, 100 ms
   "HMI_CUBA_FESTO_HMI_SENSOR_DSBG_BASTIDOR_ARRIBA_2" : Bool = PLC HMI_CUBA_FESTO.HMI_SENSOR_DSBG_BASTIDOR_ARRIBA_2, 100 ms
   "HMI_CUBA_FESTO_HMI_SENSOR_DSBG_BASTIDOR_ABAJO_2" : Bool = PLC HMI_CUBA_FESTO.HMI_SENSOR_DSBG_BASTIDOR_ABAJO_2, 100 ms
   "HMI_CUBA_FESTO_HMI_PULSADOR_SUBIR_1" : Bool = PLC HMI_CUBA_FESTO.HMI_PULSADOR_SUBIR_1, 100 ms
   "HMI_CUBA_FESTO_HMI_PULSADOR_BAJAR_1" : Bool = PLC HMI_CUBA_FESTO.HMI_PULSADOR_BAJAR_1, 100 ms
   "HMI_CUBA_FESTO_HMI_PULSADOR_SUBIR_2" : Bool = PLC HMI_CUBA_FESTO.HMI_PULSADOR_SUBIR_2, 100 ms
   "HMI_CUBA_FESTO_HMI_PULSADOR_BAJAR_2" : Bool = PLC HMI_CUBA_FESTO.HMI_PULSADOR_BAJAR_2, 100 ms
   "HMI_CUBA_FESTO_HMI_VALVULA_52_BIESTABLE_11" : Bool = PLC HMI_CUBA_FESTO.HMI_VALVULA_52_BIESTABLE_11, 100 ms
   "HMI_CUBA_FESTO_HMI_VALVULA_52_BIESTABLE_12" : Bool = PLC HMI_CUBA_FESTO.HMI_VALVULA_52_BIESTABLE_12, 100 ms
   "HMI_CUBA_FESTO_HMI_VALVULA_52_BIESTABLE_21" : Bool = PLC HMI_CUBA_FESTO.HMI_VALVULA_52_BIESTABLE_21 AT %DB1.DBX0.0, 100 ms
   "HMI_CUBA_FESTO_HMI_VALVULA_52_BIESTABLE_22" : Bool = PLC HMI_CUBA_FESTO.HMI_VALVULA_52_BIESTABLE_22 AT %DB1.DBX0.0, 100 ms
   "HMI_CUBA_FESTO_HMI_VÁLVULA_52_MONOESTABLE_1" : Bool = PLC HMI_CUBA_FESTO.HMI_VÁLVULA_52_MONOESTABLE_1 AT %DB1.DBX0.0, 100 ms
   "HMI_CUBA_FESTO_HMI_VÁLVULA_52_MONOESTABLE_2" : Bool = PLC HMI_CUBA_FESTO.HMI_VÁLVULA_52_MONOESTABLE_2 AT %DB1.DBX0.0, 100 ms
   "HMI_CUBA_FESTO_HMI_VÁLVULA_52_MONOESTABLE_3" : Bool = PLC HMI_CUBA_FESTO.HMI_VÁLVULA_52_MONOESTABLE_3 AT %DB1.DBX0.0, 100 ms
   "HMI_CUBA_FESTO_HMI_VÁLVULA_52_MONOESTABLE_4" : Bool = PLC HMI_CUBA_FESTO.HMI_VÁLVULA_52_MONOESTABLE_4 AT %DB1.DBX0.0, 100 ms
   "HMI_CUBA_FESTO_HMI_VÁLVULA_52_MONOESTABLE_5" : Bool = PLC HMI_CUBA_FESTO.HMI_VÁLVULA_52_MONOESTABLE_5 AT %DB1.DBX0.0, 100 ms
   "HMI_CUBA_FESTO_HMI_VÁLVULA_52_MONOESTABLE_6" : Bool = PLC HMI_CUBA_FESTO.HMI_VÁLVULA_52_MONOESTABLE_6 AT %DB1.DBX0.0, 100 ms
   "HMI_CUBA_FESTO_HMI_VÁLVULA_52_MONOESTABLE_7" : Bool = PLC HMI_CUBA_FESTO.HMI_VÁLVULA_52_MONOESTABLE_7 AT %DB1.DBX0.0, 100 ms
   "HMI_CUBA_FESTO_HMI_VÁLVULA_52_MONOESTABLE_8" : Bool = PLC HMI_CUBA_FESTO.HMI_VÁLVULA_52_MONOESTABLE_8 AT %DB1.DBX0.0, 100 ms
   "HMI_CUBA_FESTO_HMI_VÁLVULA_52_MONOESTABLE_9" : Bool = PLC HMI_CUBA_FESTO.HMI_VÁLVULA_52_MONOESTABLE_9 AT %DB1.DBX0.0, 100 ms
   "HMI_CUBA_FESTO_HMI_VÁLVULA_52_MONOESTABLE_10" : Bool = PLC HMI_CUBA_FESTO.HMI_VÁLVULA_52_MONOESTABLE_10 AT %DB1.DBX0.0, 100 ms
   "HMI_CUBA_FESTO_HMI_VÁLVULA_52_MONOESTABLE_11" : Bool = PLC HMI_CUBA_FESTO.HMI_VÁLVULA_52_MONOESTABLE_11 AT %DB1.DBX0.0, 100 ms
   "HMI_CUBA_FESTO_HMI_VÁLVULA_52_MONOESTABLE_12" : Bool = PLC HMI_CUBA_FESTO.HMI_VÁLVULA_52_MONOESTABLE_12 AT %DB1.DBX0.0, 100 ms
   "HMI_CUBA_FESTO_HMI_VÁLVULA_52_MONOESTABLE_13" : Bool = PLC HMI_CUBA_FESTO.HMI_VÁLVULA_52_MONOESTABLE_13 AT %DB1.DBX0.0, 100 ms
   "HMI_CUBA_FESTO_HMI_VÁLVULA_52_MONOESTABLE_14" : Bool = PLC HMI_CUBA_FESTO.HMI_VÁLVULA_52_MONOESTABLE_14 AT %DB1.DBX0.0, 100 ms
   "HMI_CUBA_FESTO_HMI_VÁLVULA_52_MONOESTABLE_15" : Bool = PLC HMI_CUBA_FESTO.HMI_VÁLVULA_52_MONOESTABLE_15 AT %DB1.DBX0.0, 100 ms
   "HMI_CUBA_FESTO_HMI_VÁLVULA_52_MONOESTABLE_16" : Bool = PLC HMI_CUBA_FESTO.HMI_VÁLVULA_52_MONOESTABLE_16 AT %DB1.DBX0.0, 100 ms
   "HMI_CUBA_FESTO_HMI_VÁLVULA_52_MONOESTABLE_17" : Bool = PLC HMI_CUBA_FESTO.HMI_VÁLVULA_52_MONOESTABLE_17 AT %DB1.DBX0.0, 100 ms
   "HMI_CUBA_FESTO_HMI_VÁLVULA_52_MONOESTABLE_18" : Bool = PLC HMI_CUBA_FESTO.HMI_VÁLVULA_52_MONOESTABLE_18 AT %DB1.DBX0.0, 100 ms
   "HMI_CUBA_FESTO_HMI_VÁLVULA_52_MONOESTABLE_19" : Bool = PLC HMI_CUBA_FESTO.HMI_VÁLVULA_52_MONOESTABLE_19 AT %DB1.DBX0.0, 100 ms